REGION Network 12: Voyage_TIME
   RUNG wire#powerrail
      Mul(in1 := "2115_VOYAGE_TIME_DAYS".VOYAGE_DAYS, in2 := 1440.0, out => "2115_VOYAGE_TIME_DAYS".VOYAGE_MINUTE)
      Mul(in1 := "2115_VOYAGE_TIME_DAYS".VOYAGE_DAYS, in2 := 24.0, out => "2115_VOYAGE_TIME_DAYS".VOYAGE_HOURS)
      Sub(in1 := "2102_TIME_CALCS_DB".TOT_SEQ_MINS, in2 := "2115_VOYAGE_TIME_DAYS".VOYAGE_MINUTE, out => "2102_TIME_CALCS_DB".Voyage_TIME_shorter_min)
      Sub(in1 := "2110_BTCS_CNTRL_DB".TOT_SEQ_HRS, in2 := "2115_VOYAGE_TIME_DAYS".VOYAGE_HOURS, out => "2102_TIME_CALCS_DB".Voyage_TIME_shorter_hours)
      Div(in1 := "2102_TIME_CALCS_DB".PRE_DWELL_MINS, in2 := 60, out => "2102_TIME_CALCS_DB".PRE_DWELL_HRS)
      { S7_Templates := "SrcType := Int"; S7_Expression := "IN1-(IN2-IN3)" } Calculate(in1 := "2102_TIME_CALCS_DB".Voyage_TIME_remaining_h, in2 := "2110_BTCS_CNTRL_DB".TOT_SEQ_HRS, in3 := "2102_TIME_CALCS_DB".PRE_DWELL_HRS, out => "2102_TIME_CALCS_DB"."PRE-DWEL HOURS REMNG")
      { S7_Templates := "SrcType := Int"; S7_Expression := "(IN1-(IN2-IN3))-(((IN4*IN5)*(IN4*IN5))/(IN4*IN5))" } Calculate(in1 := "2102_TIME_CALCS_DB".Voyage_TIME_remaining_m, in2 := "2102_TIME_CALCS_DB".TOT_SEQ_MINS, in3 := "2102_TIME_CALCS_DB".PRE_DWELL_MINS, in4 := "2102_TIME_CALCS_DB"."PRE-DWEL HOURS REMNG", in5 := 60, out => "2102_TIME_CALCS_DB"."PRE-DWEL MINS REMNG")
      { S7_Templates := "[SrcType := Int, DestType := Real]" } Convert(in := "2110_BTCS_CNTRL_DB".TOT_SEQ_HRS, out => #T_REAL)
      { S7_Templates := "SrcType := Real" } LT_Contact(in1 := "2115_VOYAGE_TIME_DAYS".VOYAGE_HOURS, in2 := #T_REAL)
      Contact( "AlwaysTRUE" )
      Coil( "2102_TIME_CALCS_DB".Voyage_TIME_invalid )
   END_RUNG
   // the same network as SCL:
   "2115_VOYAGE_TIME_DAYS".VOYAGE_MINUTE := "2115_VOYAGE_TIME_DAYS".VOYAGE_DAYS * 1440.0;
   "2115_VOYAGE_TIME_DAYS".VOYAGE_HOURS := "2115_VOYAGE_TIME_DAYS".VOYAGE_DAYS * 24.0;
   "2102_TIME_CALCS_DB".Voyage_TIME_shorter_min := "2102_TIME_CALCS_DB".TOT_SEQ_MINS - "2115_VOYAGE_TIME_DAYS".VOYAGE_MINUTE;
   "2102_TIME_CALCS_DB".Voyage_TIME_shorter_hours := "2110_BTCS_CNTRL_DB".TOT_SEQ_HRS - "2115_VOYAGE_TIME_DAYS".VOYAGE_HOURS;
   "2102_TIME_CALCS_DB".PRE_DWELL_HRS := "2102_TIME_CALCS_DB".PRE_DWELL_MINS / 60;
   "2102_TIME_CALCS_DB"."PRE-DWEL HOURS REMNG" := "2102_TIME_CALCS_DB".Voyage_TIME_remaining_h-("2110_BTCS_CNTRL_DB".TOT_SEQ_HRS-"2102_TIME_CALCS_DB".PRE_DWELL_HRS);
   "2102_TIME_CALCS_DB"."PRE-DWEL MINS REMNG" := ("2102_TIME_CALCS_DB".Voyage_TIME_remaining_m-("2102_TIME_CALCS_DB".TOT_SEQ_MINS-"2102_TIME_CALCS_DB".PRE_DWELL_MINS))-((("2102_TIME_CALCS_DB"."PRE-DWEL HOURS REMNG"*60)*("2102_TIME_CALCS_DB"."PRE-DWEL HOURS REMNG"*60))/("2102_TIME_CALCS_DB"."PRE-DWEL HOURS REMNG"*60));
   #T_REAL := INT_TO_REAL("2110_BTCS_CNTRL_DB".TOT_SEQ_HRS);
   "2102_TIME_CALCS_DB".Voyage_TIME_invalid := ("2115_VOYAGE_TIME_DAYS".VOYAGE_HOURS < #T_REAL) AND "AlwaysTRUE";
END_REGION

REGION Network 13: Caculate Time Until Treatment Required
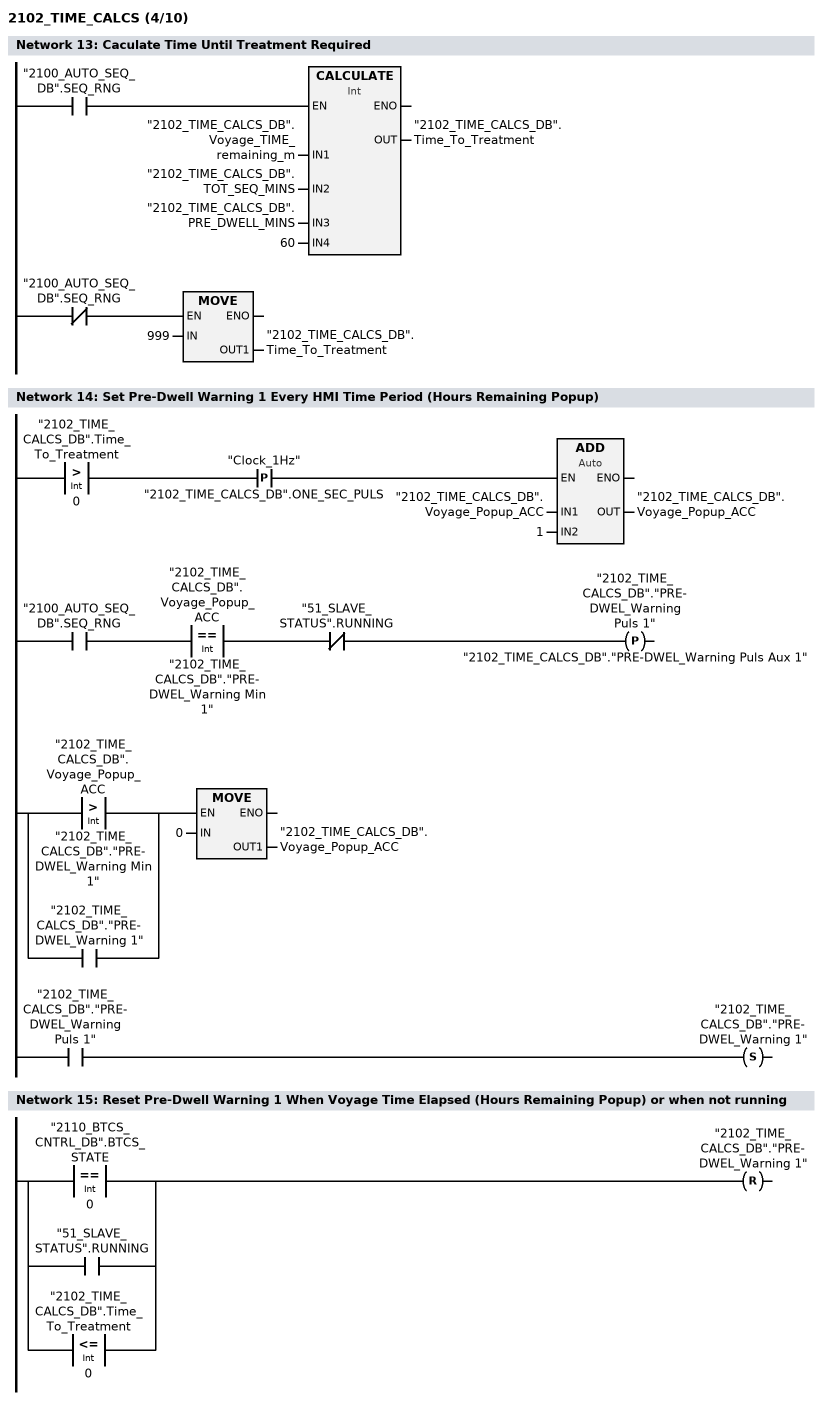
   RUNG wire#powerrail
      Contact( "2100_AUTO_SEQ_DB".SEQ_RNG )
      { S7_Templates := "SrcType := Int"; S7_Expression := "(IN1 - (IN2 - IN3)) / IN4" } Calculate(in1 := "2102_TIME_CALCS_DB".Voyage_TIME_remaining_m, in2 := "2102_TIME_CALCS_DB".TOT_SEQ_MINS, in3 := "2102_TIME_CALCS_DB".PRE_DWELL_MINS, in4 := 60, out => "2102_TIME_CALCS_DB".Time_To_Treatment)
   END_RUNG
   RUNG wire#powerrail
      I_Contact( "2100_AUTO_SEQ_DB".SEQ_RNG )
      Move(in := 999, out1 => "2102_TIME_CALCS_DB".Time_To_Treatment)
   END_RUNG
   // the same network as SCL:
   IF "2100_AUTO_SEQ_DB".SEQ_RNG THEN
       "2102_TIME_CALCS_DB".Time_To_Treatment := ("2102_TIME_CALCS_DB".Voyage_TIME_remaining_m - ("2102_TIME_CALCS_DB".TOT_SEQ_MINS - "2102_TIME_CALCS_DB".PRE_DWELL_MINS)) / 60;
   END_IF;
   IF NOT "2100_AUTO_SEQ_DB".SEQ_RNG THEN "2102_TIME_CALCS_DB".Time_To_Treatment := 999; END_IF;
END_REGION

REGION Network 14: Set Pre-Dwell Warning 1 Every HMI Time Period (Hours Remaining Popup)
   #_w1 := ("2102_TIME_CALCS_DB".Time_To_Treatment > 0) AND "Clock_1Hz" AND NOT "2102_TIME_CALCS_DB".ONE_SEC_PULS;   // rising edge of "Clock_1Hz"
   "2102_TIME_CALCS_DB".ONE_SEC_PULS := "Clock_1Hz";
   IF #_w1 THEN "2102_TIME_CALCS_DB".Voyage_Popup_ACC := "2102_TIME_CALCS_DB".Voyage_Popup_ACC + 1; END_IF;
   #_w2 := "2100_AUTO_SEQ_DB".SEQ_RNG AND ("2102_TIME_CALCS_DB".Voyage_Popup_ACC = "2102_TIME_CALCS_DB"."PRE-DWEL_Warning Min 1") AND NOT "51_SLAVE_STATUS".RUNNING;
   "2102_TIME_CALCS_DB"."PRE-DWEL_Warning Puls 1" := #_w2 AND NOT "2102_TIME_CALCS_DB"."PRE-DWEL_Warning Puls Aux 1";   // rising edge
   "2102_TIME_CALCS_DB"."PRE-DWEL_Warning Puls Aux 1" := #_w2;
   IF ("2102_TIME_CALCS_DB".Voyage_Popup_ACC > "2102_TIME_CALCS_DB"."PRE-DWEL_Warning Min 1") OR "2102_TIME_CALCS_DB"."PRE-DWEL_Warning 1" THEN
       "2102_TIME_CALCS_DB".Voyage_Popup_ACC := 0;
   END_IF;
   IF "2102_TIME_CALCS_DB"."PRE-DWEL_Warning Puls 1" THEN
       "2102_TIME_CALCS_DB"."PRE-DWEL_Warning 1" := TRUE;
   END_IF;
END_REGION

REGION Network 15: Reset Pre-Dwell Warning 1 When Voyage Time Elapsed (Hours Remaining Popup) or when not running
   RUNG wire#powerrail
      { S7_Templates := "SrcType := Int" } EQ_Contact(in1 := "2110_BTCS_CNTRL_DB".BTCS_STATE, in2 := 0)
      wire#w1
      R_Coil( "2102_TIME_CALCS_DB"."PRE-DWEL_Warning 1" )
   END_RUNG
   RUNG wire#powerrail
      Contact( "51_SLAVE_STATUS".RUNNING )
   END_RUNG wire#w1
   RUNG wire#powerrail
      { S7_Templates := "SrcType := Int" } LE_Contact(in1 := "2102_TIME_CALCS_DB".Time_To_Treatment, in2 := 0)
   END_RUNG wire#w1
   // the same network as SCL:
   IF ("2110_BTCS_CNTRL_DB".BTCS_STATE = 0) OR "51_SLAVE_STATUS".RUNNING OR ("2102_TIME_CALCS_DB".Time_To_Treatment <= 0) THEN
       "2102_TIME_CALCS_DB"."PRE-DWEL_Warning 1" := FALSE;
   END_IF;
END_REGION

REGION Network 16: Set Pre-Dwell Warning 2 When Voyage Time Elapsed (BTCS Enabled Popup) (Reset from HMI)
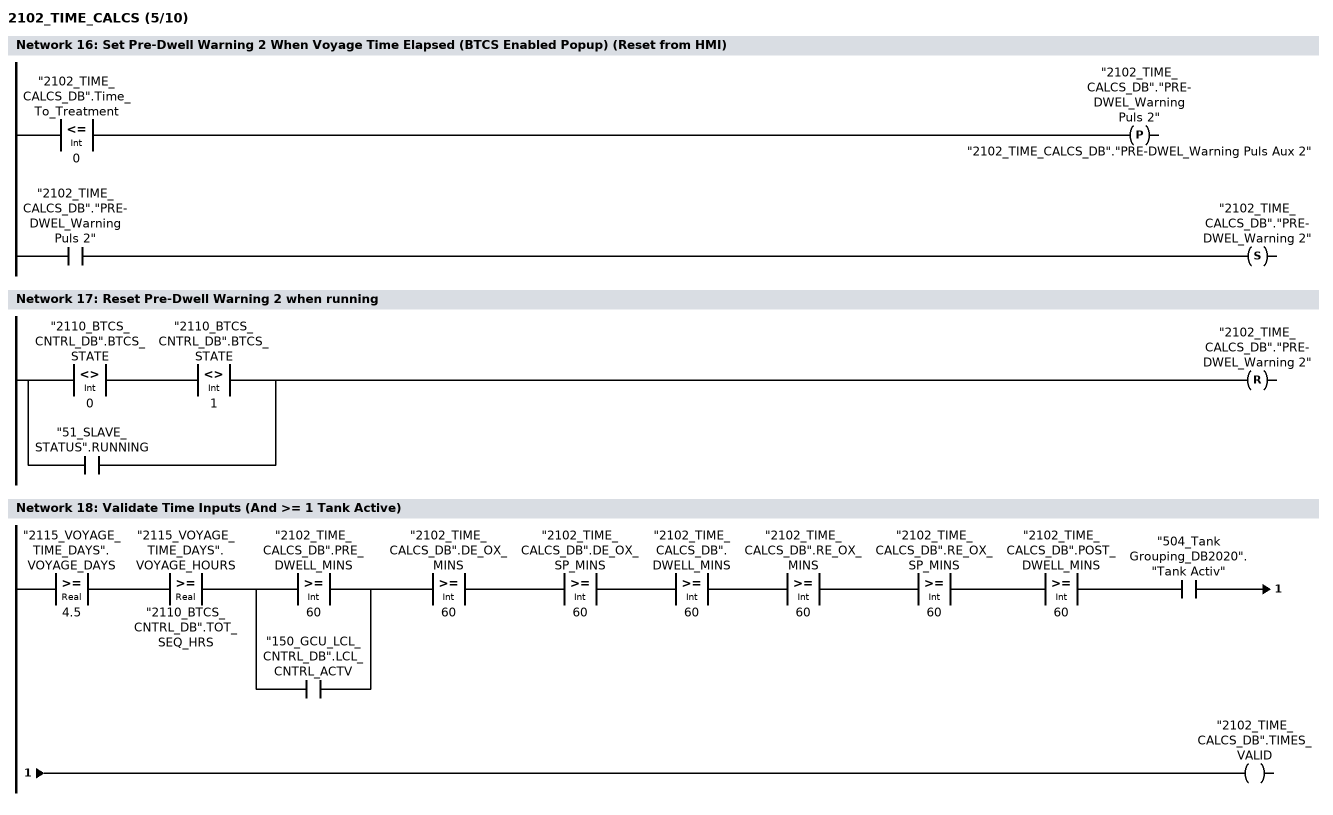
   #_w1 := "2102_TIME_CALCS_DB".Time_To_Treatment <= 0;
   "2102_TIME_CALCS_DB"."PRE-DWEL_Warning Puls 2" := #_w1 AND NOT "2102_TIME_CALCS_DB"."PRE-DWEL_Warning Puls Aux 2";   // rising edge
   "2102_TIME_CALCS_DB"."PRE-DWEL_Warning Puls Aux 2" := #_w1;
   IF "2102_TIME_CALCS_DB"."PRE-DWEL_Warning Puls 2" THEN
       "2102_TIME_CALCS_DB"."PRE-DWEL_Warning 2" := TRUE;
   END_IF;
END_REGION

REGION Network 17: Reset Pre-Dwell Warning 2 when running
   RUNG wire#powerrail
      { S7_Templates := "SrcType := Int" } NE_Contact(in1 := "2110_BTCS_CNTRL_DB".BTCS_STATE, in2 := 0)
      { S7_Templates := "SrcType := Int" } NE_Contact(in1 := "2110_BTCS_CNTRL_DB".BTCS_STATE, in2 := 1)
      wire#w1
      R_Coil( "2102_TIME_CALCS_DB"."PRE-DWEL_Warning 2" )
   END_RUNG
   RUNG wire#powerrail
      Contact( "51_SLAVE_STATUS".RUNNING )
   END_RUNG wire#w1
   // the same network as SCL:
   IF (("2110_BTCS_CNTRL_DB".BTCS_STATE <> 0) AND ("2110_BTCS_CNTRL_DB".BTCS_STATE <> 1)) OR "51_SLAVE_STATUS".RUNNING THEN
       "2102_TIME_CALCS_DB"."PRE-DWEL_Warning 2" := FALSE;
   END_IF;
END_REGION

REGION Network 18: Validate Time Inputs (And >= 1 Tank Active)
   RUNG wire#powerrail
      { S7_Templates := "SrcType := Real" } GE_Contact(in1 := "2115_VOYAGE_TIME_DAYS".VOYAGE_DAYS, in2 := 4.5)
      { S7_Templates := "SrcType := Real" } GE_Contact(in1 := "2115_VOYAGE_TIME_DAYS".VOYAGE_HOURS, in2 := "2110_BTCS_CNTRL_DB".TOT_SEQ_HRS)
      wire#w1
      { S7_Templates := "SrcType := Int" } GE_Contact(in1 := "2102_TIME_CALCS_DB".PRE_DWELL_MINS, in2 := 60)
      wire#w2
      { S7_Templates := "SrcType := Int" } GE_Contact(in1 := "2102_TIME_CALCS_DB".DE_OX_MINS, in2 := 60)
      { S7_Templates := "SrcType := Int" } GE_Contact(in1 := "2102_TIME_CALCS_DB".DE_OX_SP_MINS, in2 := 60)
      { S7_Templates := "SrcType := Int" } GE_Contact(in1 := "2102_TIME_CALCS_DB".DWELL_MINS, in2 := 60)
      { S7_Templates := "SrcType := Int" } GE_Contact(in1 := "2102_TIME_CALCS_DB".RE_OX_MINS, in2 := 60)
      { S7_Templates := "SrcType := Int" } GE_Contact(in1 := "2102_TIME_CALCS_DB".RE_OX_SP_MINS, in2 := 60)
      { S7_Templates := "SrcType := Int" } GE_Contact(in1 := "2102_TIME_CALCS_DB".POST_DWELL_MINS, in2 := 60)
      Contact( "504_Tank Grouping_DB2020"."Tank Activ" )
      Coil( "2102_TIME_CALCS_DB".TIMES_VALID )
   END_RUNG
   RUNG wire#w1
      Contact( "150_GCU_LCL_CNTRL_DB".LCL_CNTRL_ACTV )
   END_RUNG wire#w2
   // the same network as SCL:
   "2102_TIME_CALCS_DB".TIMES_VALID := ("2115_VOYAGE_TIME_DAYS".VOYAGE_DAYS >= 4.5) AND ("2115_VOYAGE_TIME_DAYS".VOYAGE_HOURS >= "2110_BTCS_CNTRL_DB".TOT_SEQ_HRS) AND (("2102_TIME_CALCS_DB".PRE_DWELL_MINS >= 60) OR "150_GCU_LCL_CNTRL_DB".LCL_CNTRL_ACTV) AND ("2102_TIME_CALCS_DB".DE_OX_MINS >= 60) AND ("2102_TIME_CALCS_DB".DE_OX_SP_MINS >= 60) AND ("2102_TIME_CALCS_DB".DWELL_MINS >= 60) AND ("2102_TIME_CALCS_DB".RE_OX_MINS >= 60) AND ("2102_TIME_CALCS_DB".RE_OX_SP_MINS >= 60) AND ("2102_TIME_CALCS_DB".POST_DWELL_MINS >= 60) AND "504_Tank Grouping_DB2020"."Tank Activ";
END_REGION

REGION Network 19: Write Values To Remaining Time
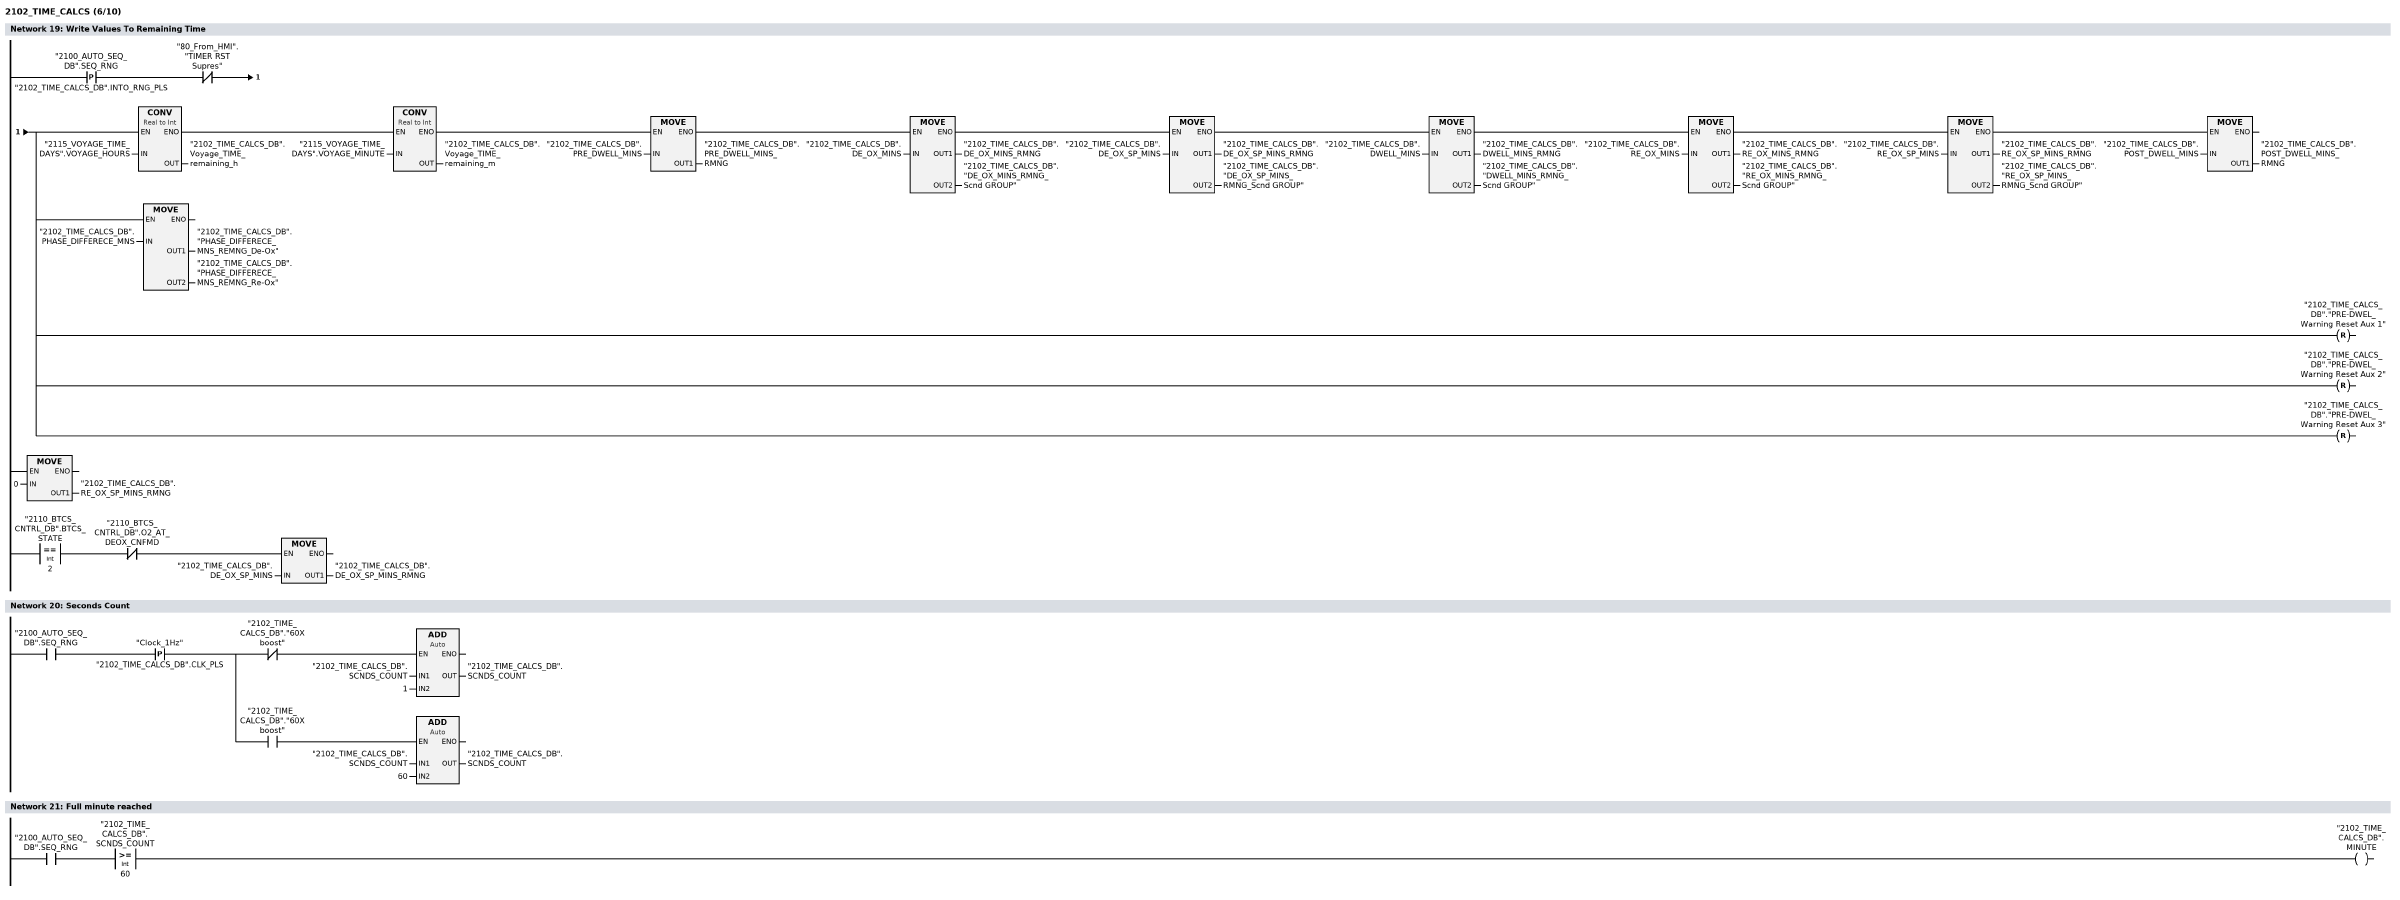
   RUNG wire#powerrail
      P_Contact(operand := "2100_AUTO_SEQ_DB".SEQ_RNG, bit := "2102_TIME_CALCS_DB".INTO_RNG_PLS)
      I_Contact( "80_From_HMI"."TIMER RST Supres" )
      wire#w1
      { S7_Templates := "[SrcType := Real, DestType := Int]" } Convert(in := "2115_VOYAGE_TIME_DAYS".VOYAGE_HOURS, out => "2102_TIME_CALCS_DB".Voyage_TIME_remaining_h)
      { S7_Templates := "[SrcType := Real, DestType := Int]" } Convert(in := "2115_VOYAGE_TIME_DAYS".VOYAGE_MINUTE, out => "2102_TIME_CALCS_DB".Voyage_TIME_remaining_m)
      Move(in := "2102_TIME_CALCS_DB".PRE_DWELL_MINS, out1 => "2102_TIME_CALCS_DB".PRE_DWELL_MINS_RMNG)
      Move(in := "2102_TIME_CALCS_DB".DE_OX_MINS, out1 => "2102_TIME_CALCS_DB".DE_OX_MINS_RMNG, out2 => "2102_TIME_CALCS_DB"."DE_OX_MINS_RMNG_Scnd GROUP")
      Move(in := "2102_TIME_CALCS_DB".DE_OX_SP_MINS, out1 => "2102_TIME_CALCS_DB".DE_OX_SP_MINS_RMNG, out2 => "2102_TIME_CALCS_DB"."DE_OX_SP_MINS_RMNG_Scnd GROUP")
      Move(in := "2102_TIME_CALCS_DB".DWELL_MINS, out1 => "2102_TIME_CALCS_DB".DWELL_MINS_RMNG, out2 => "2102_TIME_CALCS_DB"."DWELL_MINS_RMNG_Scnd GROUP")
      Move(in := "2102_TIME_CALCS_DB".RE_OX_MINS, out1 => "2102_TIME_CALCS_DB".RE_OX_MINS_RMNG, out2 => "2102_TIME_CALCS_DB"."RE_OX_MINS_RMNG_Scnd GROUP")
      Move(in := "2102_TIME_CALCS_DB".RE_OX_SP_MINS, out1 => "2102_TIME_CALCS_DB".RE_OX_SP_MINS_RMNG, out2 => "2102_TIME_CALCS_DB"."RE_OX_SP_MINS_RMNG_Scnd GROUP")
      Move(in := "2102_TIME_CALCS_DB".POST_DWELL_MINS, out1 => "2102_TIME_CALCS_DB".POST_DWELL_MINS_RMNG)
   END_RUNG
   RUNG wire#w1
      Move(in := "2102_TIME_CALCS_DB".PHASE_DIFFERECE_MNS, out1 => "2102_TIME_CALCS_DB"."PHASE_DIFFERECE_MNS_REMNG_De-Ox", out2 => "2102_TIME_CALCS_DB"."PHASE_DIFFERECE_MNS_REMNG_Re-Ox")
   END_RUNG
   RUNG wire#w1
      R_Coil( "2102_TIME_CALCS_DB"."PRE-DWEL_Warning Reset Aux 1" )
   END_RUNG
   RUNG wire#w1
      R_Coil( "2102_TIME_CALCS_DB"."PRE-DWEL_Warning Reset Aux 2" )
   END_RUNG
   RUNG wire#w1
      R_Coil( "2102_TIME_CALCS_DB"."PRE-DWEL_Warning Reset Aux 3" )
   END_RUNG
   RUNG wire#powerrail
      Move(in := 0, out1 => "2102_TIME_CALCS_DB".RE_OX_SP_MINS_RMNG)
   END_RUNG
   RUNG wire#powerrail
      { S7_Templates := "SrcType := Int" } EQ_Contact(in1 := "2110_BTCS_CNTRL_DB".BTCS_STATE, in2 := 2)
      I_Contact( "2110_BTCS_CNTRL_DB".O2_AT_DEOX_CNFMD )
      Move(in := "2102_TIME_CALCS_DB".DE_OX_SP_MINS, out1 => "2102_TIME_CALCS_DB".DE_OX_SP_MINS_RMNG)
   END_RUNG
   // the same network as SCL:
   #_w1 := "2100_AUTO_SEQ_DB".SEQ_RNG AND NOT "2102_TIME_CALCS_DB".INTO_RNG_PLS;   // rising edge of "2100_AUTO_SEQ_DB".SEQ_RNG
   "2102_TIME_CALCS_DB".INTO_RNG_PLS := "2100_AUTO_SEQ_DB".SEQ_RNG;
   IF #_w1 AND NOT "80_From_HMI"."TIMER RST Supres" THEN
       "2102_TIME_CALCS_DB".Voyage_TIME_remaining_h := REAL_TO_INT("2115_VOYAGE_TIME_DAYS".VOYAGE_HOURS);
       "2102_TIME_CALCS_DB".Voyage_TIME_remaining_m := REAL_TO_INT("2115_VOYAGE_TIME_DAYS".VOYAGE_MINUTE);
       "2102_TIME_CALCS_DB".PRE_DWELL_MINS_RMNG := "2102_TIME_CALCS_DB".PRE_DWELL_MINS;
       "2102_TIME_CALCS_DB".DE_OX_MINS_RMNG := "2102_TIME_CALCS_DB".DE_OX_MINS;
       "2102_TIME_CALCS_DB"."DE_OX_MINS_RMNG_Scnd GROUP" := "2102_TIME_CALCS_DB".DE_OX_MINS;
       "2102_TIME_CALCS_DB".DE_OX_SP_MINS_RMNG := "2102_TIME_CALCS_DB".DE_OX_SP_MINS;
       "2102_TIME_CALCS_DB"."DE_OX_SP_MINS_RMNG_Scnd GROUP" := "2102_TIME_CALCS_DB".DE_OX_SP_MINS;
       "2102_TIME_CALCS_DB".DWELL_MINS_RMNG := "2102_TIME_CALCS_DB".DWELL_MINS;
       "2102_TIME_CALCS_DB"."DWELL_MINS_RMNG_Scnd GROUP" := "2102_TIME_CALCS_DB".DWELL_MINS;
       "2102_TIME_CALCS_DB".RE_OX_MINS_RMNG := "2102_TIME_CALCS_DB".RE_OX_MINS;
       "2102_TIME_CALCS_DB"."RE_OX_MINS_RMNG_Scnd GROUP" := "2102_TIME_CALCS_DB".RE_OX_MINS;
       "2102_TIME_CALCS_DB".RE_OX_SP_MINS_RMNG := "2102_TIME_CALCS_DB".RE_OX_SP_MINS;
       "2102_TIME_CALCS_DB"."RE_OX_SP_MINS_RMNG_Scnd GROUP" := "2102_TIME_CALCS_DB".RE_OX_SP_MINS;
       "2102_TIME_CALCS_DB".POST_DWELL_MINS_RMNG := "2102_TIME_CALCS_DB".POST_DWELL_MINS;
       "2102_TIME_CALCS_DB"."PHASE_DIFFERECE_MNS_REMNG_De-Ox" := "2102_TIME_CALCS_DB".PHASE_DIFFERECE_MNS;
       "2102_TIME_CALCS_DB"."PHASE_DIFFERECE_MNS_REMNG_Re-Ox" := "2102_TIME_CALCS_DB".PHASE_DIFFERECE_MNS;
       "2102_TIME_CALCS_DB"."PRE-DWEL_Warning Reset Aux 1" := FALSE;
       "2102_TIME_CALCS_DB"."PRE-DWEL_Warning Reset Aux 2" := FALSE;
       "2102_TIME_CALCS_DB"."PRE-DWEL_Warning Reset Aux 3" := FALSE;
   END_IF;
   "2102_TIME_CALCS_DB".RE_OX_SP_MINS_RMNG := 0;
   IF ("2110_BTCS_CNTRL_DB".BTCS_STATE = 2) AND NOT "2110_BTCS_CNTRL_DB".O2_AT_DEOX_CNFMD THEN
       "2102_TIME_CALCS_DB".DE_OX_SP_MINS_RMNG := "2102_TIME_CALCS_DB".DE_OX_SP_MINS;
   END_IF;
END_REGION

REGION Network 20: Seconds Count
   RUNG wire#powerrail
      Contact( "2100_AUTO_SEQ_DB".SEQ_RNG )
      P_Contact(operand := "Clock_1Hz", bit := "2102_TIME_CALCS_DB".CLK_PLS)
      wire#w1
      I_Contact( "2102_TIME_CALCS_DB"."60X boost" )
      Add(in1 := "2102_TIME_CALCS_DB".SCNDS_COUNT, in2 := 1, out => "2102_TIME_CALCS_DB".SCNDS_COUNT)
   END_RUNG
   RUNG wire#w1
      Contact( "2102_TIME_CALCS_DB"."60X boost" )
      Add(in1 := "2102_TIME_CALCS_DB".SCNDS_COUNT, in2 := 60, out => "2102_TIME_CALCS_DB".SCNDS_COUNT)
   END_RUNG
   // the same network as SCL:
   #_w1 := "2100_AUTO_SEQ_DB".SEQ_RNG AND "Clock_1Hz" AND NOT "2102_TIME_CALCS_DB".CLK_PLS;   // rising edge of "Clock_1Hz"
   "2102_TIME_CALCS_DB".CLK_PLS := "Clock_1Hz";
   IF #_w1 AND NOT "2102_TIME_CALCS_DB"."60X boost" THEN
       "2102_TIME_CALCS_DB".SCNDS_COUNT := "2102_TIME_CALCS_DB".SCNDS_COUNT + 1;
   END_IF;
   IF #_w1 AND "2102_TIME_CALCS_DB"."60X boost" THEN
       "2102_TIME_CALCS_DB".SCNDS_COUNT := "2102_TIME_CALCS_DB".SCNDS_COUNT + 60;
   END_IF;
END_REGION

REGION Network 21: Full minute reached
   RUNG wire#powerrail
      Contact( "2100_AUTO_SEQ_DB".SEQ_RNG )
      { S7_Templates := "SrcType := Int" } GE_Contact(in1 := "2102_TIME_CALCS_DB".SCNDS_COUNT, in2 := 60)
      Coil( "2102_TIME_CALCS_DB".MINUTE )
   END_RUNG
   // the same network as SCL:
   "2102_TIME_CALCS_DB".MINUTE := "2100_AUTO_SEQ_DB".SEQ_RNG AND ("2102_TIME_CALCS_DB".SCNDS_COUNT >= 60);
END_REGION

REGION Network 22: Count Downs
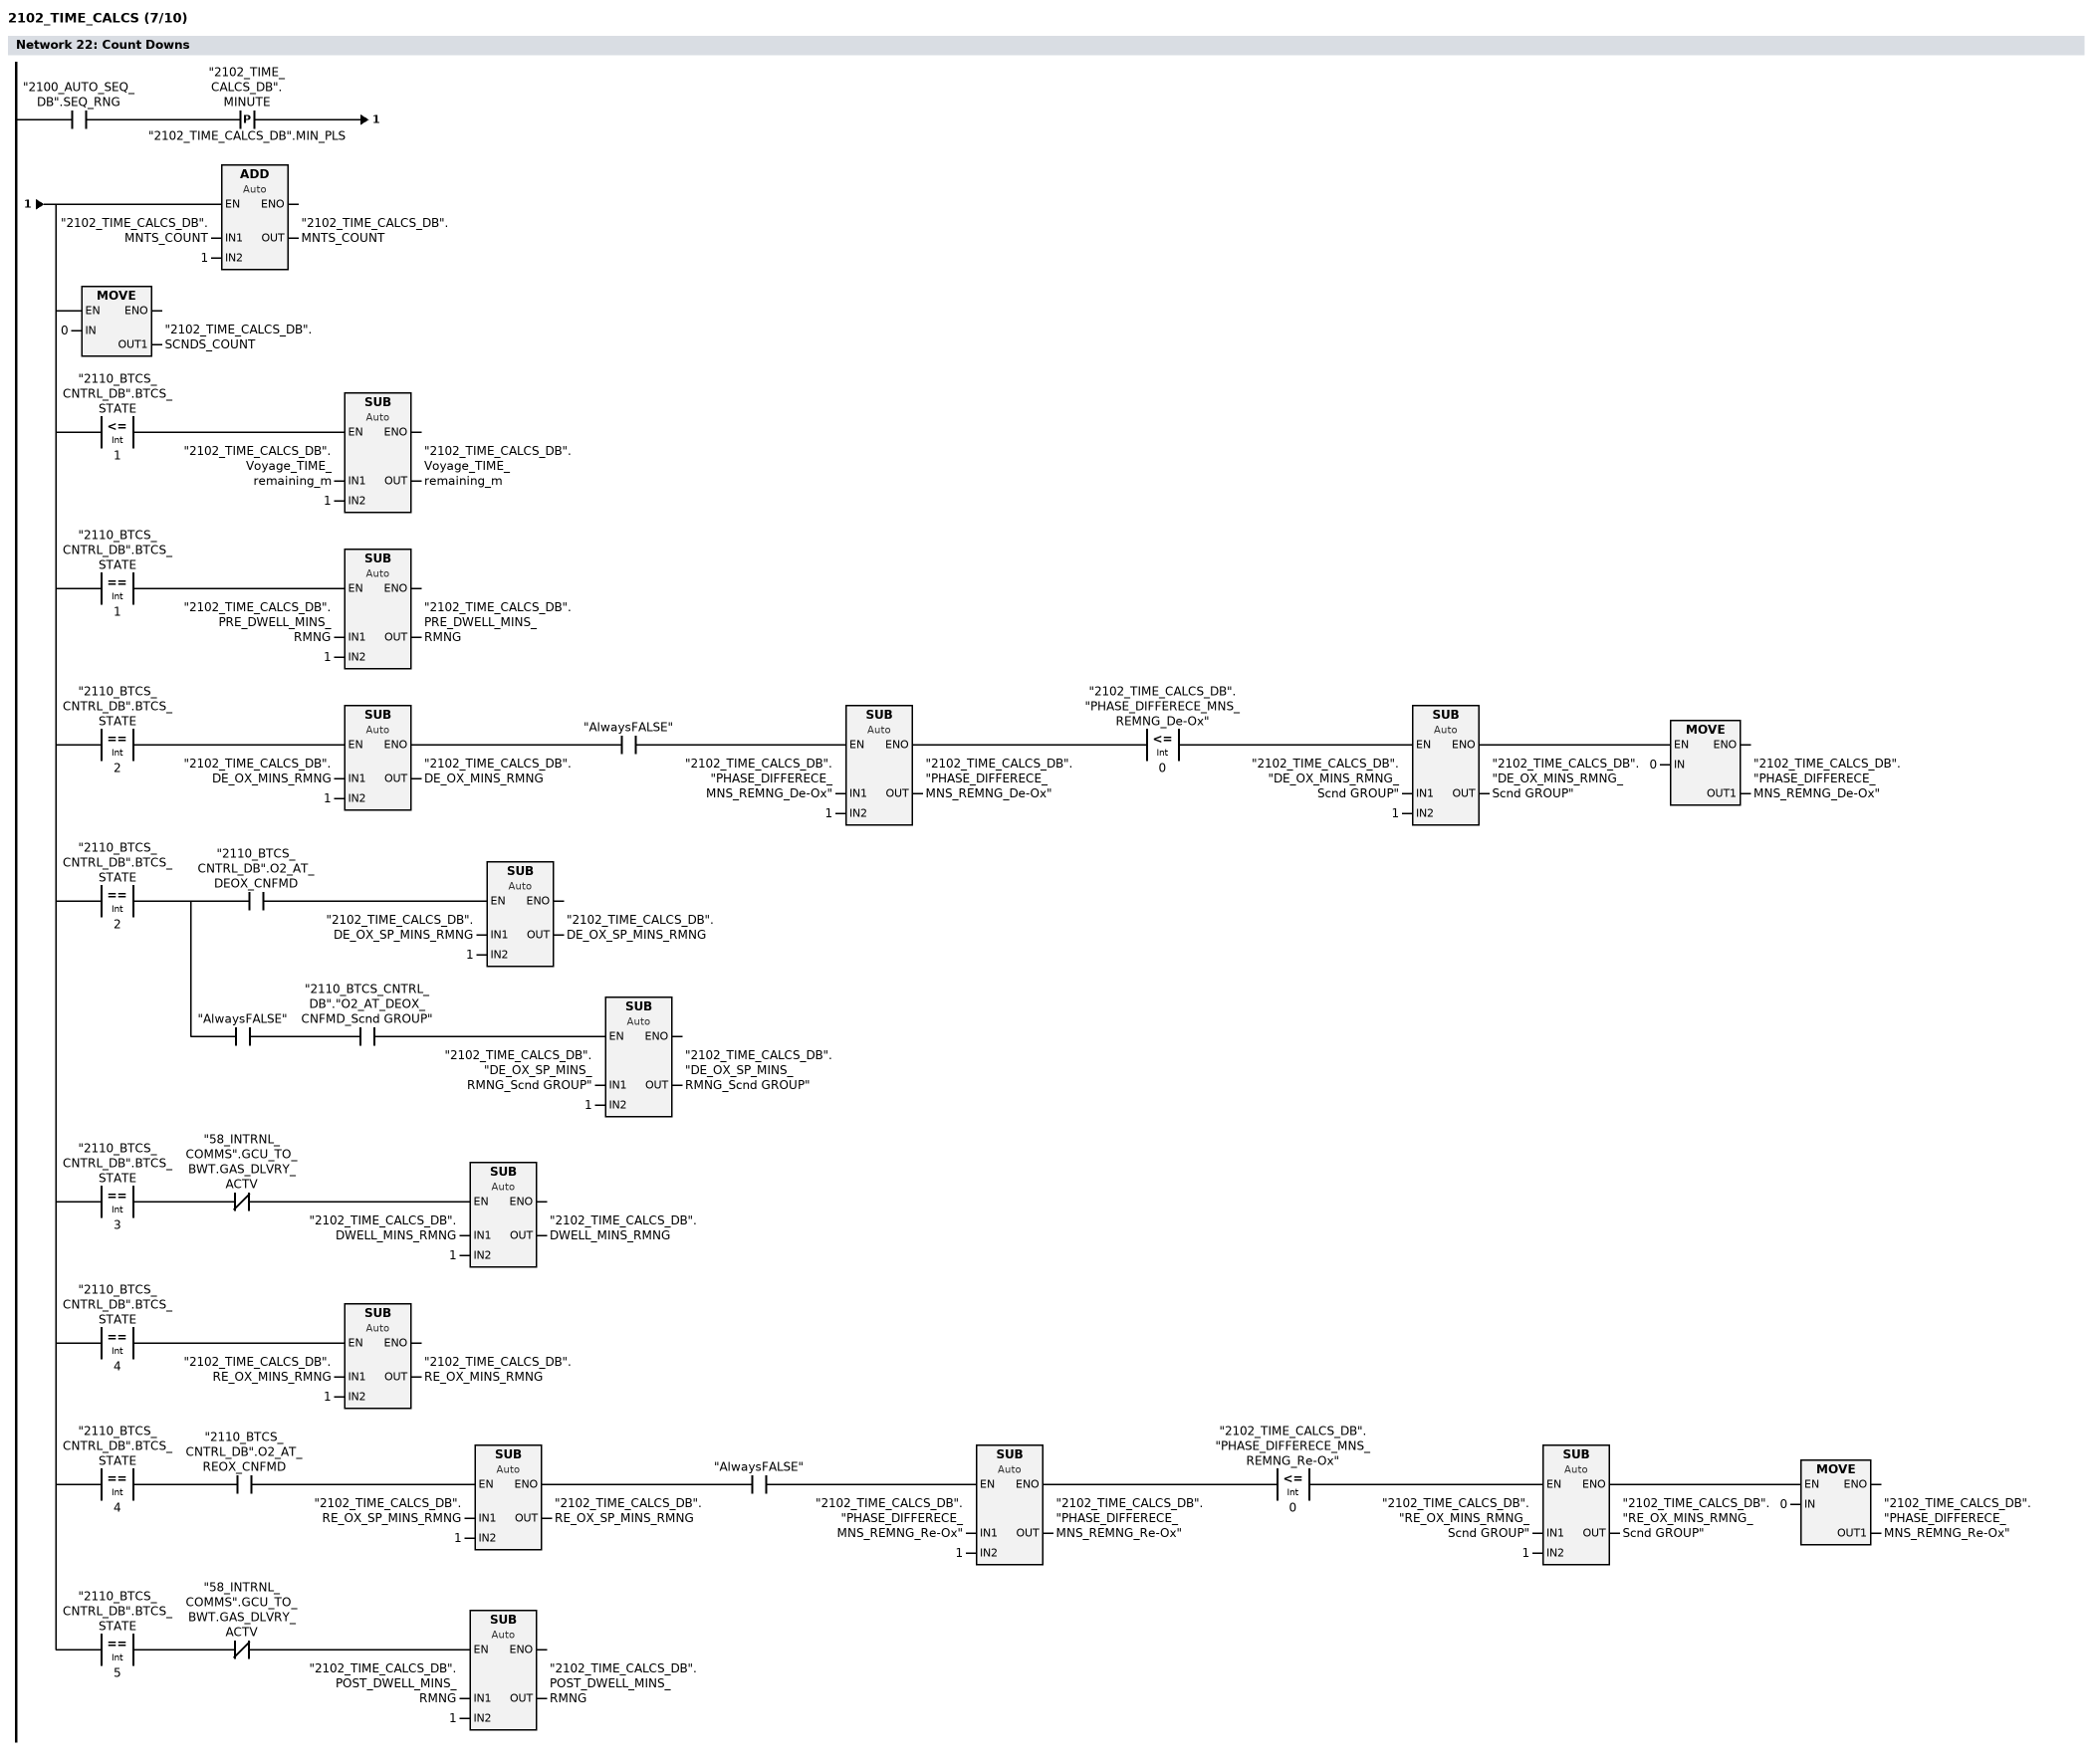
   RUNG wire#powerrail
      Contact( "2100_AUTO_SEQ_DB".SEQ_RNG )
      P_Contact(operand := "2102_TIME_CALCS_DB".MINUTE, bit := "2102_TIME_CALCS_DB".MIN_PLS)
      wire#w1
      Add(in1 := "2102_TIME_CALCS_DB".MNTS_COUNT, in2 := 1, out => "2102_TIME_CALCS_DB".MNTS_COUNT)
   END_RUNG
   RUNG wire#w1
      Move(in := 0, out1 => "2102_TIME_CALCS_DB".SCNDS_COUNT)
   END_RUNG
   RUNG wire#w1
      { S7_Templates := "SrcType := Int" } LE_Contact(in1 := "2110_BTCS_CNTRL_DB".BTCS_STATE, in2 := 1)
      Sub(in1 := "2102_TIME_CALCS_DB".Voyage_TIME_remaining_m, in2 := 1, out => "2102_TIME_CALCS_DB".Voyage_TIME_remaining_m)
   END_RUNG
   RUNG wire#w1
      { S7_Templates := "SrcType := Int" } EQ_Contact(in1 := "2110_BTCS_CNTRL_DB".BTCS_STATE, in2 := 1)
      Sub(in1 := "2102_TIME_CALCS_DB".PRE_DWELL_MINS_RMNG, in2 := 1, out => "2102_TIME_CALCS_DB".PRE_DWELL_MINS_RMNG)
   END_RUNG
   RUNG wire#w1
      { S7_Templates := "SrcType := Int" } EQ_Contact(in1 := "2110_BTCS_CNTRL_DB".BTCS_STATE, in2 := 2)
      Sub(in1 := "2102_TIME_CALCS_DB".DE_OX_MINS_RMNG, in2 := 1, out => "2102_TIME_CALCS_DB".DE_OX_MINS_RMNG)
      Contact( "AlwaysFALSE" )
      Sub(in1 := "2102_TIME_CALCS_DB"."PHASE_DIFFERECE_MNS_REMNG_De-Ox", in2 := 1, out => "2102_TIME_CALCS_DB"."PHASE_DIFFERECE_MNS_REMNG_De-Ox")
      { S7_Templates := "SrcType := Int" } LE_Contact(in1 := "2102_TIME_CALCS_DB"."PHASE_DIFFERECE_MNS_REMNG_De-Ox", in2 := 0)
      Sub(in1 := "2102_TIME_CALCS_DB"."DE_OX_MINS_RMNG_Scnd GROUP", in2 := 1, out => "2102_TIME_CALCS_DB"."DE_OX_MINS_RMNG_Scnd GROUP")
      Move(in := 0, out1 => "2102_TIME_CALCS_DB"."PHASE_DIFFERECE_MNS_REMNG_De-Ox")
   END_RUNG
   RUNG wire#w1
      { S7_Templates := "SrcType := Int" } EQ_Contact(in1 := "2110_BTCS_CNTRL_DB".BTCS_STATE, in2 := 2)
      wire#w2
      Contact( "2110_BTCS_CNTRL_DB".O2_AT_DEOX_CNFMD )
      Sub(in1 := "2102_TIME_CALCS_DB".DE_OX_SP_MINS_RMNG, in2 := 1, out => "2102_TIME_CALCS_DB".DE_OX_SP_MINS_RMNG)
   END_RUNG
   RUNG wire#w2
      Contact( "AlwaysFALSE" )
      Contact( "2110_BTCS_CNTRL_DB"."O2_AT_DEOX_CNFMD_Scnd GROUP" )
      Sub(in1 := "2102_TIME_CALCS_DB"."DE_OX_SP_MINS_RMNG_Scnd GROUP", in2 := 1, out => "2102_TIME_CALCS_DB"."DE_OX_SP_MINS_RMNG_Scnd GROUP")
   END_RUNG
   RUNG wire#w1
      { S7_Templates := "SrcType := Int" } EQ_Contact(in1 := "2110_BTCS_CNTRL_DB".BTCS_STATE, in2 := 3)
      I_Contact( "58_INTRNL_COMMS".GCU_TO_BWT.GAS_DLVRY_ACTV )
      Sub(in1 := "2102_TIME_CALCS_DB".DWELL_MINS_RMNG, in2 := 1, out => "2102_TIME_CALCS_DB".DWELL_MINS_RMNG)
   END_RUNG
   RUNG wire#w1
      { S7_Templates := "SrcType := Int" } EQ_Contact(in1 := "2110_BTCS_CNTRL_DB".BTCS_STATE, in2 := 4)
      Sub(in1 := "2102_TIME_CALCS_DB".RE_OX_MINS_RMNG, in2 := 1, out => "2102_TIME_CALCS_DB".RE_OX_MINS_RMNG)
   END_RUNG
   RUNG wire#w1
      { S7_Templates := "SrcType := Int" } EQ_Contact(in1 := "2110_BTCS_CNTRL_DB".BTCS_STATE, in2 := 4)
      Contact( "2110_BTCS_CNTRL_DB".O2_AT_REOX_CNFMD )
      Sub(in1 := "2102_TIME_CALCS_DB".RE_OX_SP_MINS_RMNG, in2 := 1, out => "2102_TIME_CALCS_DB".RE_OX_SP_MINS_RMNG)
      Contact( "AlwaysFALSE" )
      Sub(in1 := "2102_TIME_CALCS_DB"."PHASE_DIFFERECE_MNS_REMNG_Re-Ox", in2 := 1, out => "2102_TIME_CALCS_DB"."PHASE_DIFFERECE_MNS_REMNG_Re-Ox")
      { S7_Templates := "SrcType := Int" } LE_Contact(in1 := "2102_TIME_CALCS_DB"."PHASE_DIFFERECE_MNS_REMNG_Re-Ox", in2 := 0)
      Sub(in1 := "2102_TIME_CALCS_DB"."RE_OX_MINS_RMNG_Scnd GROUP", in2 := 1, out => "2102_TIME_CALCS_DB"."RE_OX_MINS_RMNG_Scnd GROUP")
      Move(in := 0, out1 => "2102_TIME_CALCS_DB"."PHASE_DIFFERECE_MNS_REMNG_Re-Ox")
   END_RUNG
   RUNG wire#w1
      { S7_Templates := "SrcType := Int" } EQ_Contact(in1 := "2110_BTCS_CNTRL_DB".BTCS_STATE, in2 := 5)
      I_Contact( "58_INTRNL_COMMS".GCU_TO_BWT.GAS_DLVRY_ACTV )
      Sub(in1 := "2102_TIME_CALCS_DB".POST_DWELL_MINS_RMNG, in2 := 1, out => "2102_TIME_CALCS_DB".POST_DWELL_MINS_RMNG)
   END_RUNG
   // the same network as SCL:
   #_w1 := "2100_AUTO_SEQ_DB".SEQ_RNG AND "2102_TIME_CALCS_DB".MINUTE AND NOT "2102_TIME_CALCS_DB".MIN_PLS;   // rising edge of "2102_TIME_CALCS_DB".MINUTE
   "2102_TIME_CALCS_DB".MIN_PLS := "2102_TIME_CALCS_DB".MINUTE;
   IF #_w1 THEN
       "2102_TIME_CALCS_DB".MNTS_COUNT := "2102_TIME_CALCS_DB".MNTS_COUNT + 1;
       "2102_TIME_CALCS_DB".SCNDS_COUNT := 0;
   END_IF;
   IF #_w1 AND ("2110_BTCS_CNTRL_DB".BTCS_STATE <= 1) THEN
       "2102_TIME_CALCS_DB".Voyage_TIME_remaining_m := "2102_TIME_CALCS_DB".Voyage_TIME_remaining_m - 1;
   END_IF;
   IF #_w1 AND ("2110_BTCS_CNTRL_DB".BTCS_STATE = 1) THEN
       "2102_TIME_CALCS_DB".PRE_DWELL_MINS_RMNG := "2102_TIME_CALCS_DB".PRE_DWELL_MINS_RMNG - 1;
   END_IF;
   #_w2 := #_w1 AND ("2110_BTCS_CNTRL_DB".BTCS_STATE = 2);
   IF #_w2 THEN "2102_TIME_CALCS_DB".DE_OX_MINS_RMNG := "2102_TIME_CALCS_DB".DE_OX_MINS_RMNG - 1; END_IF;
   #_w3 := #_w2 AND "AlwaysFALSE";
   IF #_w3 THEN
       "2102_TIME_CALCS_DB"."PHASE_DIFFERECE_MNS_REMNG_De-Ox" := "2102_TIME_CALCS_DB"."PHASE_DIFFERECE_MNS_REMNG_De-Ox" - 1;
   END_IF;
   IF #_w3 AND ("2102_TIME_CALCS_DB"."PHASE_DIFFERECE_MNS_REMNG_De-Ox" <= 0) THEN
       "2102_TIME_CALCS_DB"."DE_OX_MINS_RMNG_Scnd GROUP" := "2102_TIME_CALCS_DB"."DE_OX_MINS_RMNG_Scnd GROUP" - 1;
       "2102_TIME_CALCS_DB"."PHASE_DIFFERECE_MNS_REMNG_De-Ox" := 0;
   END_IF;
   #_w4 := #_w1 AND ("2110_BTCS_CNTRL_DB".BTCS_STATE = 2);
   IF #_w4 AND "2110_BTCS_CNTRL_DB".O2_AT_DEOX_CNFMD THEN
       "2102_TIME_CALCS_DB".DE_OX_SP_MINS_RMNG := "2102_TIME_CALCS_DB".DE_OX_SP_MINS_RMNG - 1;
   END_IF;
   IF #_w4 AND "AlwaysFALSE" AND "2110_BTCS_CNTRL_DB"."O2_AT_DEOX_CNFMD_Scnd GROUP" THEN
       "2102_TIME_CALCS_DB"."DE_OX_SP_MINS_RMNG_Scnd GROUP" := "2102_TIME_CALCS_DB"."DE_OX_SP_MINS_RMNG_Scnd GROUP" - 1;
   END_IF;
   IF #_w1 AND ("2110_BTCS_CNTRL_DB".BTCS_STATE = 3) AND NOT "58_INTRNL_COMMS".GCU_TO_BWT.GAS_DLVRY_ACTV THEN
       "2102_TIME_CALCS_DB".DWELL_MINS_RMNG := "2102_TIME_CALCS_DB".DWELL_MINS_RMNG - 1;
   END_IF;
   IF #_w1 AND ("2110_BTCS_CNTRL_DB".BTCS_STATE = 4) THEN
       "2102_TIME_CALCS_DB".RE_OX_MINS_RMNG := "2102_TIME_CALCS_DB".RE_OX_MINS_RMNG - 1;
   END_IF;
   #_w5 := #_w1 AND ("2110_BTCS_CNTRL_DB".BTCS_STATE = 4) AND "2110_BTCS_CNTRL_DB".O2_AT_REOX_CNFMD;
   IF #_w5 THEN
       "2102_TIME_CALCS_DB".RE_OX_SP_MINS_RMNG := "2102_TIME_CALCS_DB".RE_OX_SP_MINS_RMNG - 1;
   END_IF;
   #_w6 := #_w5 AND "AlwaysFALSE";
   IF #_w6 THEN
       "2102_TIME_CALCS_DB"."PHASE_DIFFERECE_MNS_REMNG_Re-Ox" := "2102_TIME_CALCS_DB"."PHASE_DIFFERECE_MNS_REMNG_Re-Ox" - 1;
   END_IF;
   IF #_w6 AND ("2102_TIME_CALCS_DB"."PHASE_DIFFERECE_MNS_REMNG_Re-Ox" <= 0) THEN
       "2102_TIME_CALCS_DB"."RE_OX_MINS_RMNG_Scnd GROUP" := "2102_TIME_CALCS_DB"."RE_OX_MINS_RMNG_Scnd GROUP" - 1;
       "2102_TIME_CALCS_DB"."PHASE_DIFFERECE_MNS_REMNG_Re-Ox" := 0;
   END_IF;
   IF #_w1 AND ("2110_BTCS_CNTRL_DB".BTCS_STATE = 5) AND NOT "58_INTRNL_COMMS".GCU_TO_BWT.GAS_DLVRY_ACTV THEN
       "2102_TIME_CALCS_DB".POST_DWELL_MINS_RMNG := "2102_TIME_CALCS_DB".POST_DWELL_MINS_RMNG - 1;
   END_IF;
END_REGION

REGION Network 23: Full hour reached
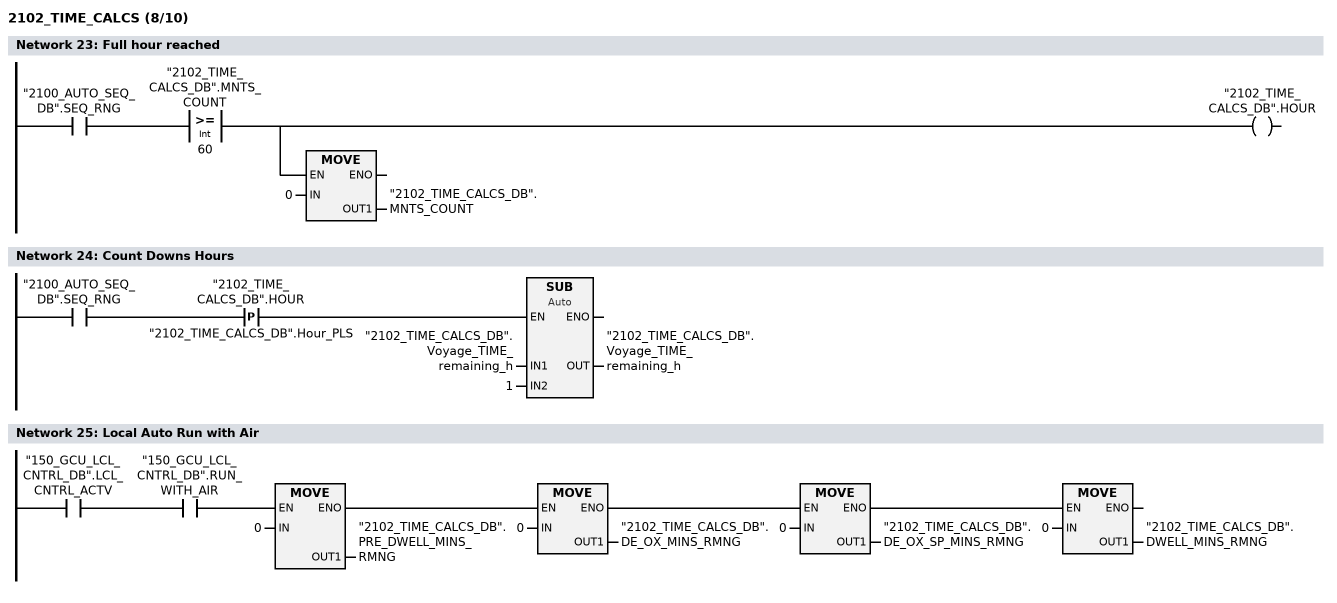
   RUNG wire#powerrail
      Contact( "2100_AUTO_SEQ_DB".SEQ_RNG )
      { S7_Templates := "SrcType := Int" } GE_Contact(in1 := "2102_TIME_CALCS_DB".MNTS_COUNT, in2 := 60)
      wire#w1
      Coil( "2102_TIME_CALCS_DB".HOUR )
   END_RUNG
   RUNG wire#w1
      Move(in := 0, out1 => "2102_TIME_CALCS_DB".MNTS_COUNT)
   END_RUNG
   // the same network as SCL:
   "2102_TIME_CALCS_DB".HOUR := "2100_AUTO_SEQ_DB".SEQ_RNG AND ("2102_TIME_CALCS_DB".MNTS_COUNT >= 60);
   IF "2102_TIME_CALCS_DB".HOUR THEN "2102_TIME_CALCS_DB".MNTS_COUNT := 0; END_IF;
END_REGION

REGION Network 24: Count Downs Hours
   RUNG wire#powerrail
      Contact( "2100_AUTO_SEQ_DB".SEQ_RNG )
      P_Contact(operand := "2102_TIME_CALCS_DB".HOUR, bit := "2102_TIME_CALCS_DB".Hour_PLS)
      Sub(in1 := "2102_TIME_CALCS_DB".Voyage_TIME_remaining_h, in2 := 1, out => "2102_TIME_CALCS_DB".Voyage_TIME_remaining_h)
   END_RUNG
   // the same network as SCL:
   #_w1 := "2100_AUTO_SEQ_DB".SEQ_RNG AND "2102_TIME_CALCS_DB".HOUR AND NOT "2102_TIME_CALCS_DB".Hour_PLS;   // rising edge of "2102_TIME_CALCS_DB".HOUR
   "2102_TIME_CALCS_DB".Hour_PLS := "2102_TIME_CALCS_DB".HOUR;
   IF #_w1 THEN
       "2102_TIME_CALCS_DB".Voyage_TIME_remaining_h := "2102_TIME_CALCS_DB".Voyage_TIME_remaining_h - 1;
   END_IF;
END_REGION

REGION Network 25: Local Auto Run with Air
   RUNG wire#powerrail
      Contact( "150_GCU_LCL_CNTRL_DB".LCL_CNTRL_ACTV )
      Contact( "150_GCU_LCL_CNTRL_DB".RUN_WITH_AIR )
      Move(in := 0, out1 => "2102_TIME_CALCS_DB".PRE_DWELL_MINS_RMNG)
      Move(in := 0, out1 => "2102_TIME_CALCS_DB".DE_OX_MINS_RMNG)
      Move(in := 0, out1 => "2102_TIME_CALCS_DB".DE_OX_SP_MINS_RMNG)
      Move(in := 0, out1 => "2102_TIME_CALCS_DB".DWELL_MINS_RMNG)
   END_RUNG
   // the same network as SCL:
   IF "150_GCU_LCL_CNTRL_DB".LCL_CNTRL_ACTV AND "150_GCU_LCL_CNTRL_DB".RUN_WITH_AIR THEN
       "2102_TIME_CALCS_DB".PRE_DWELL_MINS_RMNG := 0;
       "2102_TIME_CALCS_DB".DE_OX_MINS_RMNG := 0;
       "2102_TIME_CALCS_DB".DE_OX_SP_MINS_RMNG := 0;
       "2102_TIME_CALCS_DB".DWELL_MINS_RMNG := 0;
   END_IF;
END_REGION

